HMI tags "ProNet Configuration"
   "PN_Mixinghead_Send" : Bool = PLC PN_Mixinghead.Send AT %DB1006.DBX4.0, 1 s
   "PN_Mixinghead_Mixinghead{0}_Digital_Address" : Int = PLC PN_Mixinghead.Mixinghead[0].Digital.Address AT %DB1006.DBW80, 1 s
      on ChangeValue: SetBit("PN_Mixinghead_Mixinghead{0}_Digital_Zeiten_Request"); SetBit("PN_Mixinghead_Mixinghead{0}_Digital_Zeiten_2_Request"); SetBit("PN_Mixinghead_Mixinghead{0}_Digital_GeneralParameters_Request")
   "PN_Mixinghead_Mixinghead{0}_Digital_Zeiten_Request" : Bool = PLC PN_Mixinghead.Mixinghead[0].Digital.Zeiten.Request AT %DB1006.DBX90.0, 1 s
   "PN_Mixinghead_Mixinghead{0}_Digital_Zeiten_Data_ÜberwachungszeitÖffnen" : Real = PLC PN_Mixinghead.Mixinghead[0].Digital.Zeiten.Data.ÜberwachungszeitÖffnen AT %DB1006.DBD92, 1 s
      on ChangeValue: SetBit("PN_Mixinghead_Mixinghead{0}_Digital_Zeiten_Request")
   "PN_Mixinghead_Mixinghead{0}_Digital_GeneralParameters_Data_MischkopfKanal" : Byte = PLC PN_Mixinghead.Mixinghead[0].Digital.GeneralParameters.Data.MischkopfKanal AT %DB1006.DBB89, 1 s
      on ChangeValue: SetBit("PN_Mixinghead_Mixinghead{0}_Digital_GeneralParameters_Request")
   "PN_Mixinghead_Mixinghead{0}_Digital_GeneralParameters_Request" : Bool = PLC PN_Mixinghead.Mixinghead[0].Digital.GeneralParameters.Request AT %DB1006.DBX84.0, 1 s
   "PN_Mixinghead_Mixinghead{0}_Digital_Active" : Bool = PLC PN_Mixinghead.Mixinghead[0].Digital.Active AT %DB1006.DBX82.0, 1 s
      on ChangeValue: SetBit("PN_Mixinghead_Mixinghead{0}_Digital_Zeiten_Request"); SetBit("PN_Mixinghead_Mixinghead{0}_Digital_Zeiten_2_Request"); SetBit("PN_Mixinghead_Mixinghead{0}_Digital_GeneralParameters_Request")
   "PN_Mixinghead_Mixinghead{0}_Digital_Zeiten_Data_ÜberwachungszeitSchließen" : Real = PLC PN_Mixinghead.Mixinghead[0].Digital.Zeiten.Data.ÜberwachungszeitSchließen AT %DB1006.DBD96, 1 s
      on ChangeValue: SetBit("PN_Mixinghead_Mixinghead{0}_Digital_Zeiten_Request")
   "PN_Mixinghead_Mixinghead{0}_Digital_Zeiten_Data_ErlaubtePrellzeit" : Real = PLC PN_Mixinghead.Mixinghead[0].Digital.Zeiten.Data.ErlaubtePrellzeit AT %DB1006.DBD100, 1 s
      on ChangeValue: SetBit("PN_Mixinghead_Mixinghead{0}_Digital_Zeiten_Request")
   "PN_Mixinghead_Mixinghead{0}_Digital_GeneralParameters_Data_Ventilausgang" : Byte = PLC PN_Mixinghead.Mixinghead[0].Digital.GeneralParameters.Data.Ventilausgang AT %DB1006.DBB88, 1 s
      on ChangeValue: SetBit("PN_Mixinghead_Mixinghead{0}_Digital_GeneralParameters_Request")
   "PN_Mixinghead_Mixinghead{0}_Digital_GeneralParameters_Data_EingangskanalMK_Ini" : Byte = PLC PN_Mixinghead.Mixinghead[0].Digital.GeneralParameters.Data.EingangskanalMK_Ini AT %DB1006.DBB86, 1 s
      on ChangeValue: SetBit("PN_Mixinghead_Mixinghead{0}_Digital_GeneralParameters_Request")
   "PN_Mixinghead_Mixinghead{0}_Digital_GeneralParameters_Data_EingangskanalFreigabe" : Byte = PLC PN_Mixinghead.Mixinghead[0].Digital.GeneralParameters.Data.EingangskanalFreigabe AT %DB1006.DBB87, 1 s
      on ChangeValue: SetBit("PN_Mixinghead_Mixinghead{0}_Digital_GeneralParameters_Request")
   "PN_Mixinghead_Mixinghead{0}_Digital_Zeiten_2_Request" : Bool = PLC PN_Mixinghead.Mixinghead[0].Digital.Zeiten_2.Request AT %DB1006.DBX104.0, 1 s
   "PN_Mixinghead_Mixinghead{0}_Digital_Zeiten_2_Data_Verzögerungszeit_HW_Freigabe" : Real = PLC PN_Mixinghead.Mixinghead[0].Digital.Zeiten_2.Data.Verzögerungszeit_HW_Freigabe AT %DB1006.DBD106, 1 s
      on ChangeValue: SetBit("PN_Mixinghead_Mixinghead{0}_Digital_Zeiten_2_Request")
   "PN_Mixinghead_SetIndex" : Int = PLC PN_Mixinghead.SetIndex AT %DB1006.DBW0, 1 s
   "PN_Mixinghead_Mixinghead{0}_ReinigungskolbenDigital_Active" : Bool = PLC PN_Mixinghead.Mixinghead[0].ReinigungskolbenDigital.Active AT %DB1006.DBX112.0, 1 s
      on ChangeValue: SetBit("PN_Mixinghead_Mixinghead{0}_ReinigungskolbenDigital_Zeiten_Request"); SetBit("PN_Mixinghead_Mixinghead{0}_ReinigungskolbenDigital_GeneralParameters_Request")
   "PN_Mixinghead_Mixinghead{0}_ReinigungskolbenDigital_GeneralParameters_Request" : Bool = PLC PN_Mixinghead.Mixinghead[0].ReinigungskolbenDigital.GeneralParameters.Request AT %DB1006.DBX114.0, 1 s
   "PN_Mixinghead_Mixinghead{0}_ReinigungskolbenDigital_GeneralParameters_Data_EingangskanalRK_Ini" : Byte = PLC PN_Mixinghead.Mixinghead[0].ReinigungskolbenDigital.GeneralParameters.Data.EingangskanalRK_Ini AT %DB1006.DBB116, 1 s
      on ChangeValue: SetBit("PN_Mixinghead_Mixinghead{0}_ReinigungskolbenDigital_GeneralParameters_Request")
   "PN_Mixinghead_Mixinghead{0}_ReinigungskolbenDigital_GeneralParameters_Data_AusgangRKVentil" : Byte = PLC PN_Mixinghead.Mixinghead[0].ReinigungskolbenDigital.GeneralParameters.Data.AusgangRKVentil AT %DB1006.DBB117, 1 s
      on ChangeValue: SetBit("PN_Mixinghead_Mixinghead{0}_ReinigungskolbenDigital_GeneralParameters_Request")
   "PN_Mixinghead_Mixinghead{0}_ReinigungskolbenDigital_GeneralParameters_Data_MischkopfKanal" : Byte = PLC PN_Mixinghead.Mixinghead[0].ReinigungskolbenDigital.GeneralParameters.Data.MischkopfKanal AT %DB1006.DBB118, 1 s
      on ChangeValue: SetBit("PN_Mixinghead_Mixinghead{0}_ReinigungskolbenDigital_GeneralParameters_Request")
   "PN_Mixinghead_Mixinghead{0}_ReinigungskolbenDigital_Address" : Int = PLC PN_Mixinghead.Mixinghead[0].ReinigungskolbenDigital.Address AT %DB1006.DBW110, 1 s
      on ChangeValue: SetBit("PN_Mixinghead_Mixinghead{0}_Digital_Zeiten_Request"); SetBit("PN_Mixinghead_Mixinghead{0}_Digital_Zeiten_2_Request"); SetBit("PN_Mixinghead_Mixinghead{0}_Digital_GeneralParameters_Request")
   "PN_Mixinghead_Mixinghead{0}_ReinigungskolbenDigital_Zeiten_Data_ÜberwachungszeitVorfahren" : Real = PLC PN_Mixinghead.Mixinghead[0].ReinigungskolbenDigital.Zeiten.Data.ÜberwachungszeitVorfahren AT %DB1006.DBD122, 1 s
      on ChangeValue: SetBit("PN_Mixinghead_Mixinghead{0}_ReinigungskolbenDigital_Zeiten_Request")
   "PN_Mixinghead_Mixinghead{0}_ReinigungskolbenDigital_Zeiten_Data_ÜberwachungszeitRückfahren" : Real = PLC PN_Mixinghead.Mixinghead[0].ReinigungskolbenDigital.Zeiten.Data.ÜberwachungszeitRückfahren AT %DB1006.DBD126, 1 s
      on ChangeValue: SetBit("PN_Mixinghead_Mixinghead{0}_ReinigungskolbenDigital_Zeiten_Request")
   "PN_Mixinghead_Mixinghead{0}_ReinigungskolbenDigital_Zeiten_Request" : Bool = PLC PN_Mixinghead.Mixinghead[0].ReinigungskolbenDigital.Zeiten.Request AT %DB1006.DBX120.0, 1 s
   "PN_Mixinghead_Mixinghead{0}_ReinigungskolbenDigital_Zeiten_Data_ErlaubtePrellzeit" : Real = PLC PN_Mixinghead.Mixinghead[0].ReinigungskolbenDigital.Zeiten.Data.ErlaubtePrellzeit AT %DB1006.DBD130, 1 s
      on ChangeValue: SetBit("PN_Mixinghead_Mixinghead{0}_ReinigungskolbenDigital_Zeiten_Request")
   "PN_Mixinghead_Mixinghead{0}_ReinigungskolbenDigital_Zeiten_Data_WartezeitVorne" : Real = PLC PN_Mixinghead.Mixinghead[0].ReinigungskolbenDigital.Zeiten.Data.WartezeitVorne AT %DB1006.DBD134, 1 s
      on ChangeValue: SetBit("PN_Mixinghead_Mixinghead{0}_ReinigungskolbenDigital_Zeiten_Request")
   "PN_Mixinghead_Mixinghead{0}_ReinigungskolbenDigital_Zeiten_Data_VerzögerungNachSchuss" : Real = PLC PN_Mixinghead.Mixinghead[0].ReinigungskolbenDigital.Zeiten.Data.VerzögerungNachSchuss AT %DB1006.DBD138, 1 s
      on ChangeValue: SetBit("PN_Mixinghead_Mixinghead{0}_ReinigungskolbenDigital_Zeiten_Request")
   "PN_AI_Send" : Bool = PLC PN_AI.Send AT %DB1002.DBX4.0, 1 s
   "PN_AI_Module{0}_AI8_Address" : Int = PLC PN_AI.Module[0].AI8.Address AT %DB1002.DBW6, 1 s
      on ChangeValue: SetBit("PN_AI_Send"); SetBit("PN_AI_Module{0}_AI8_X14_0_Request")
   "PN_AI_Module{0}_AI8_Active" : Bool = PLC PN_AI.Module[0].AI8.Active AT %DB1002.DBX8.0, 1 s
      on ChangeValue: SetBit("PN_AI_Send"); SetBit("PN_AI_Module{0}_AI8_X14_0_Request")
   "PN_AI_Module{0}_AI8_X14_0_Data_Data[1]_Betriebsart" : Byte = PLC PN_AI.Module[0].AI8.X14_0.Data."Data[1]".Betriebsart AT %DB1002.DBB12, 1 s
      on ChangeValue: SetBit("PN_AI_Send"); SetBit("PN_AI_Module{0}_AI8_X14_0_Request")
   "PN_AI_Module{0}_AI8_X14_0_Data_Data[2]_Betriebsart" : Byte = PLC PN_AI.Module[0].AI8.X14_0.Data."Data[2]".Betriebsart AT %DB1002.DBB20, 1 s
      on ChangeValue: SetBit("PN_AI_Send"); SetBit("PN_AI_Module{0}_AI8_X14_0_Request")
   "PN_AI_Module{0}_AI8_X14_0_Data_Data[1]_Bereichsuntergrenze" : Int = PLC PN_AI.Module[0].AI8.X14_0.Data."Data[1]".Bereichsuntergrenze AT %DB1002.DBW16, 1 s
      on ChangeValue: SetBit("PN_AI_Send"); SetBit("PN_AI_Module{0}_AI8_X14_0_Request")
   "PN_AI_Module{0}_AI8_X14_0_Data_Data[1]_Bereichsobergrenze" : Int = PLC PN_AI.Module[0].AI8.X14_0.Data."Data[1]".Bereichsobergrenze AT %DB1002.DBW14, 1 s
      on ChangeValue: SetBit("PN_AI_Send"); SetBit("PN_AI_Module{0}_AI8_X14_0_Request")
   "PN_AI_Module{0}_AI8_X14_0_Data_Data[1]_Mittelwertzeit" : Int = PLC PN_AI.Module[0].AI8.X14_0.Data."Data[1]".Mittelwertzeit AT %DB1002.DBW18, 1 s
      on ChangeValue: SetBit("PN_AI_Send"); SetBit("PN_AI_Module{0}_AI8_X14_0_Request")
   "PN_AI_Module{0}_AI8_X14_0_Data_Data[2]_Bereichsobergrenze" : Int = PLC PN_AI.Module[0].AI8.X14_0.Data."Data[2]".Bereichsobergrenze AT %DB1002.DBW22, 1 s
      on ChangeValue: SetBit("PN_AI_Send"); SetBit("PN_AI_Module{0}_AI8_X14_0_Request")
   "PN_AI_Module{0}_AI8_X14_0_Data_Data[2]_Bereichsuntergrenze" : Int = PLC PN_AI.Module[0].AI8.X14_0.Data."Data[2]".Bereichsuntergrenze AT %DB1002.DBW24, 1 s
      on ChangeValue: SetBit("PN_AI_Send"); SetBit("PN_AI_Module{0}_AI8_X14_0_Request")
   "PN_AI_Module{0}_AI8_X14_0_Data_Data[2]_Mittelwertzeit" : Int = PLC PN_AI.Module[0].AI8.X14_0.Data."Data[2]".Mittelwertzeit AT %DB1002.DBW26, 1 s
      on ChangeValue: SetBit("PN_AI_Send"); SetBit("PN_AI_Module{0}_AI8_X14_0_Request")
   "PN_AI_Module{0}_AI8_X14_0_Data_Data[3]_Betriebsart" : Byte = PLC PN_AI.Module[0].AI8.X14_0.Data."Data[3]".Betriebsart AT %DB1002.DBB28, 1 s
      on ChangeValue: SetBit("PN_AI_Send"); SetBit("PN_AI_Module{0}_AI8_X14_0_Request")
   "PN_Mixinghead_Mixinghead{0}_DüseBypass{6}_Zeiten_Request" : Bool = PLC PN_Mixinghead.Mixinghead[0].DüseBypass[6].Zeiten.Request AT %DB1006.DBX458.0, 1 s
      on ChangeValue: SetBit("PN_AI_Send"); SetBit("PN_AI_Module{0}_AI8_X14_0_Request")
   "PN_AI_Module{0}_AI8_X14_0_Data_Data[3]_Bereichsuntergrenze" : Int = PLC PN_AI.Module[0].AI8.X14_0.Data."Data[3]".Bereichsuntergrenze AT %DB1002.DBW32, 1 s
      on ChangeValue: SetBit("PN_AI_Send"); SetBit("PN_AI_Module{0}_AI8_X14_0_Request")
   "PN_AI_Module{0}_AI8_X14_0_Data_Data[3]_Mittelwertzeit" : Int = PLC PN_AI.Module[0].AI8.X14_0.Data."Data[3]".Mittelwertzeit AT %DB1002.DBW34, 1 s
      on ChangeValue: SetBit("PN_AI_Send"); SetBit("PN_AI_Module{0}_AI8_X14_0_Request")
   "PN_AI_Module{0}_AI8_X14_0_Data_Data[4]_Betriebsart" : Byte = PLC PN_AI.Module[0].AI8.X14_0.Data."Data[4]".Betriebsart AT %DB1002.DBB36, 1 s
      on ChangeValue: SetBit("PN_AI_Send"); SetBit("PN_AI_Module{0}_AI8_X14_0_Request")
   "PN_AI_Module{0}_AI8_X14_0_Data_Data[4]_Bereichsobergrenze" : Int = PLC PN_AI.Module[0].AI8.X14_0.Data."Data[4]".Bereichsobergrenze AT %DB1002.DBW38, 1 s
      on ChangeValue: SetBit("PN_AI_Send"); SetBit("PN_AI_Module{0}_AI8_X14_0_Request")
   "PN_AI_Module{0}_AI8_X14_0_Data_Data[4]_Bereichsuntergrenze" : Int = PLC PN_AI.Module[0].AI8.X14_0.Data."Data[4]".Bereichsuntergrenze AT %DB1002.DBW40, 1 s
      on ChangeValue: SetBit("PN_AI_Send"); SetBit("PN_AI_Module{0}_AI8_X14_0_Request")
   "PN_AI_Module{0}_AI8_X14_0_Data_Data[4]_Mittelwertzeit" : Int = PLC PN_AI.Module[0].AI8.X14_0.Data."Data[4]".Mittelwertzeit AT %DB1002.DBW42, 1 s
      on ChangeValue: SetBit("PN_AI_Send"); SetBit("PN_AI_Module{0}_AI8_X14_0_Request")
   "PN_AI_Module{0}_AI8_X14_0_Data_Data[5]_Betriebsart" : Byte = PLC PN_AI.Module[0].AI8.X14_0.Data."Data[5]".Betriebsart AT %DB1002.DBB44, 1 s
      on ChangeValue: SetBit("PN_AI_Send"); SetBit("PN_AI_Module{0}_AI8_X14_0_Request")
   "PN_AI_Module{0}_AI8_X14_0_Data_Data[5]_Bereichsobergrenze" : Int = PLC PN_AI.Module[0].AI8.X14_0.Data."Data[5]".Bereichsobergrenze AT %DB1002.DBW46, 1 s
      on ChangeValue: SetBit("PN_AI_Send"); SetBit("PN_AI_Module{0}_AI8_X14_0_Request")
   "PN_AI_Module{0}_AI8_X14_0_Data_Data[5]_Bereichsuntergrenze" : Int = PLC PN_AI.Module[0].AI8.X14_0.Data."Data[5]".Bereichsuntergrenze AT %DB1002.DBW48, 1 s
      on ChangeValue: SetBit("PN_AI_Send"); SetBit("PN_AI_Module{0}_AI8_X14_0_Request")
   "PN_AI_Module{0}_AI8_X14_0_Data_Data[5]_Mittelwertzeit" : Int = PLC PN_AI.Module[0].AI8.X14_0.Data."Data[5]".Mittelwertzeit AT %DB1002.DBW50, 1 s
      on ChangeValue: SetBit("PN_AI_Send"); SetBit("PN_AI_Module{0}_AI8_X14_0_Request")
   "PN_AI_Module{0}_AI8_X14_0_Data_Data[6]_Betriebsart" : Byte = PLC PN_AI.Module[0].AI8.X14_0.Data."Data[6]".Betriebsart AT %DB1002.DBB52, 1 s
      on ChangeValue: SetBit("PN_AI_Send"); SetBit("PN_AI_Module{0}_AI8_X14_0_Request")
   "PN_AI_Module{0}_AI8_X14_0_Data_Data[6]_Bereichsobergrenze" : Int = PLC PN_AI.Module[0].AI8.X14_0.Data."Data[6]".Bereichsobergrenze AT %DB1002.DBW54, 1 s
      on ChangeValue: SetBit("PN_AI_Send"); SetBit("PN_AI_Module{0}_AI8_X14_0_Request")
   "PN_AI_Module{0}_AI8_X14_0_Data_Data[6]_Bereichsuntergrenze" : Int = PLC PN_AI.Module[0].AI8.X14_0.Data."Data[6]".Bereichsuntergrenze AT %DB1002.DBW56, 1 s
      on ChangeValue: SetBit("PN_AI_Send"); SetBit("PN_AI_Module{0}_AI8_X14_0_Request")
   "PN_AI_Module{0}_AI8_X14_0_Data_Data[6]_Mittelwertzeit" : Int = PLC PN_AI.Module[0].AI8.X14_0.Data."Data[6]".Mittelwertzeit AT %DB1002.DBW58, 1 s
      on ChangeValue: SetBit("PN_AI_Send"); SetBit("PN_AI_Module{0}_AI8_X14_0_Request")
   "PN_AI_Module{0}_AI8_X14_0_Data_Data[7]_Betriebsart" : Byte = PLC PN_AI.Module[0].AI8.X14_0.Data."Data[7]".Betriebsart AT %DB1002.DBB60, 1 s
      on ChangeValue: SetBit("PN_AI_Send"); SetBit("PN_AI_Module{0}_AI8_X14_0_Request")
   "PN_AI_Module{0}_AI8_X14_0_Data_Data[7]_Bereichsobergrenze" : Int = PLC PN_AI.Module[0].AI8.X14_0.Data."Data[7]".Bereichsobergrenze AT %DB1002.DBW62, 1 s
      on ChangeValue: SetBit("PN_AI_Send"); SetBit("PN_AI_Module{0}_AI8_X14_0_Request")
   "PN_AI_Module{0}_AI8_X14_0_Data_Data[7]_Bereichsuntergrenze" : Int = PLC PN_AI.Module[0].AI8.X14_0.Data."Data[7]".Bereichsuntergrenze AT %DB1002.DBW64, 1 s
      on ChangeValue: SetBit("PN_AI_Send"); SetBit("PN_AI_Module{0}_AI8_X14_0_Request")
   "PN_AI_Module{0}_AI8_X14_0_Data_Data[7]_Mittelwertzeit" : Int = PLC PN_AI.Module[0].AI8.X14_0.Data."Data[7]".Mittelwertzeit AT %DB1002.DBW66, 1 s
      on ChangeValue: SetBit("PN_AI_Send"); SetBit("PN_AI_Module{0}_AI8_X14_0_Request")
   "PN_AI_Module{0}_AI8_X14_0_Data_Data[8]_Betriebsart" : Byte = PLC PN_AI.Module[0].AI8.X14_0.Data."Data[8]".Betriebsart AT %DB1002.DBB68, 1 s
      on ChangeValue: SetBit("PN_AI_Send"); SetBit("PN_AI_Module{0}_AI8_X14_0_Request")
   "PN_AI_Module{0}_AI8_X14_0_Data_Data[8]_Bereichsobergrenze" : Int = PLC PN_AI.Module[0].AI8.X14_0.Data."Data[8]".Bereichsobergrenze AT %DB1002.DBW70, 1 s
      on ChangeValue: SetBit("PN_AI_Send"); SetBit("PN_AI_Module{0}_AI8_X14_0_Request")
   "PN_AI_Module{0}_AI8_X14_0_Data_Data[8]_Bereichsuntergrenze" : Int = PLC PN_AI.Module[0].AI8.X14_0.Data."Data[8]".Bereichsuntergrenze AT %DB1002.DBW72, 1 s
      on ChangeValue: SetBit("PN_AI_Send"); SetBit("PN_AI_Module{0}_AI8_X14_0_Request")
   "PN_AI_Module{0}_AI8_X14_0_Data_Data[8]_Mittelwertzeit" : Int = PLC PN_AI.Module[0].AI8.X14_0.Data."Data[8]".Mittelwertzeit AT %DB1002.DBW74, 1 s
      on ChangeValue: SetBit("PN_AI_Send"); SetBit("PN_AI_Module{0}_AI8_X14_0_Request")
   "PN_AI_Module{0}_AI8_X14_0_Request" : Bool = PLC PN_AI.Module[0].AI8.X14_0.Request AT %DB1002.DBX10.0, 1 s
   "PN_AI_SetIndex" : Int = PLC PN_AI.SetIndex AT %DB1002.DBW0, 1 s
      on ChangeValue: SetBit("PN_AI_Send")
   "PN_AI_Module{0}_AIResistive_8_Address" : Int = PLC PN_AI.Module[0].AIResistive_8.Address AT %DB1002.DBW76, 1 s
      on ChangeValue: SetBit("PN_AI_Send"); SetBit("PN_AI_Module{0}_AIResistive_8_TemperatureInput_Request")
   "PN_AI_Module{0}_AIResistive_8_TemperatureInput_Request" : Bool = PLC PN_AI.Module[0].AIResistive_8.TemperatureInput.Request AT %DB1002.DBX80.0, 1 s
      on ChangeValue: SetBit("PN_AI_Send")
   "PN_AI_Module{0}_AIResistive_8_Active" : Bool = PLC PN_AI.Module[0].AIResistive_8.Active AT %DB1002.DBX78.0, 1 s
      on ChangeValue: SetBit("PN_AI_Send")
   "PN_AI_Module{0}_AIResistive_8_TemperatureInput_Data{1}_Mittelwertzeit" : Int = PLC PN_AI.Module[0].AIResistive_8.TemperatureInput.Data[1].Mittelwertzeit AT %DB1002.DBW82, 1 s
      on ChangeValue: SetBit("PN_AI_Send"); SetBit("PN_AI_Module{0}_AIResistive_8_TemperatureInput_Request")
   "PN_AI_Module{0}_AIResistive_8_TemperatureInput_Data{1}_ErsatzwertDrahtbruch" : Int = PLC PN_AI.Module[0].AIResistive_8.TemperatureInput.Data[1].ErsatzwertDrahtbruch AT %DB1002.DBW84, 1 s
      on ChangeValue: SetBit("PN_AI_Send"); SetBit("PN_AI_Module{0}_AIResistive_8_TemperatureInput_Request")
   "PN_AI_Module{0}_AIResistive_8_TemperatureInput_Data{1}_Einheit" : Byte = PLC PN_AI.Module[0].AIResistive_8.TemperatureInput.Data[1].Einheit AT %DB1002.DBB86, 1 s
      on ChangeValue: SetBit("PN_AI_Send"); SetBit("PN_AI_Module{0}_AIResistive_8_TemperatureInput_Request")
   "PN_AI_Module{0}_AIResistive_8_TemperatureInput_Data{2}_Mittelwertzeit" : Int = PLC PN_AI.Module[0].AIResistive_8.TemperatureInput.Data[2].Mittelwertzeit AT %DB1002.DBW88, 1 s
      on ChangeValue: SetBit("PN_AI_Send"); SetBit("PN_AI_Module{0}_AIResistive_8_TemperatureInput_Request")
   "PN_AI_Module{0}_AIResistive_8_TemperatureInput_Data{2}_ErsatzwertDrahtbruch" : Int = PLC PN_AI.Module[0].AIResistive_8.TemperatureInput.Data[2].ErsatzwertDrahtbruch AT %DB1002.DBW90, 1 s
      on ChangeValue: SetBit("PN_AI_Send"); SetBit("PN_AI_Module{0}_AIResistive_8_TemperatureInput_Request")
   "PN_AI_Module{0}_AIResistive_8_TemperatureInput_Data{2}_Einheit" : Byte = PLC PN_AI.Module[0].AIResistive_8.TemperatureInput.Data[2].Einheit AT %DB1002.DBB92, 1 s
      on ChangeValue: SetBit("PN_AI_Send"); SetBit("PN_AI_Module{0}_AIResistive_8_TemperatureInput_Request")
   "PN_AI_Module{0}_AIResistive_8_TemperatureInput_Data{3}_Mittelwertzeit" : Int = PLC PN_AI.Module[0].AIResistive_8.TemperatureInput.Data[3].Mittelwertzeit AT %DB1002.DBW94, 1 s
      on ChangeValue: SetBit("PN_AI_Send"); SetBit("PN_AI_Module{0}_AIResistive_8_TemperatureInput_Request")
   "PN_AI_Module{0}_AIResistive_8_TemperatureInput_Data{3}_ErsatzwertDrahtbruch" : Int = PLC PN_AI.Module[0].AIResistive_8.TemperatureInput.Data[3].ErsatzwertDrahtbruch AT %DB1002.DBW96, 1 s
      on ChangeValue: SetBit("PN_AI_Send"); SetBit("PN_AI_Module{0}_AIResistive_8_TemperatureInput_Request")
   "PN_AI_Module{0}_AIResistive_8_TemperatureInput_Data{3}_Einheit" : Byte = PLC PN_AI.Module[0].AIResistive_8.TemperatureInput.Data[3].Einheit AT %DB1002.DBB98, 1 s
      on ChangeValue: SetBit("PN_AI_Send"); SetBit("PN_AI_Module{0}_AIResistive_8_TemperatureInput_Request")
   "PN_AI_Module{0}_AIResistive_8_TemperatureInput_Data{4}_Mittelwertzeit" : Int = PLC PN_AI.Module[0].AIResistive_8.TemperatureInput.Data[4].Mittelwertzeit AT %DB1002.DBW100, 1 s
      on ChangeValue: SetBit("PN_AI_Send"); SetBit("PN_AI_Module{0}_AIResistive_8_TemperatureInput_Request")
   "PN_AI_Module{0}_AIResistive_8_TemperatureInput_Data{4}_ErsatzwertDrahtbruch" : Int = PLC PN_AI.Module[0].AIResistive_8.TemperatureInput.Data[4].ErsatzwertDrahtbruch AT %DB1002.DBW102, 1 s
      on ChangeValue: SetBit("PN_AI_Send"); SetBit("PN_AI_Module{0}_AIResistive_8_TemperatureInput_Request")
   "PN_AI_Module{0}_AIResistive_8_TemperatureInput_Data{4}_Einheit" : Byte = PLC PN_AI.Module[0].AIResistive_8.TemperatureInput.Data[4].Einheit AT %DB1002.DBB104, 1 s
      on ChangeValue: SetBit("PN_AI_Send"); SetBit("PN_AI_Module{0}_AIResistive_8_TemperatureInput_Request")
   "PN_AI_Module{0}_AIResistive_8_TemperatureInput_Data{5}_Mittelwertzeit" : Int = PLC PN_AI.Module[0].AIResistive_8.TemperatureInput.Data[5].Mittelwertzeit AT %DB1002.DBW106, 1 s
      on ChangeValue: SetBit("PN_AI_Send"); SetBit("PN_AI_Module{0}_AIResistive_8_TemperatureInput_Request")
   "PN_AI_Module{0}_AIResistive_8_TemperatureInput_Data{5}_ErsatzwertDrahtbruch" : Int = PLC PN_AI.Module[0].AIResistive_8.TemperatureInput.Data[5].ErsatzwertDrahtbruch AT %DB1002.DBW108, 1 s
      on ChangeValue: SetBit("PN_AI_Send"); SetBit("PN_AI_Module{0}_AIResistive_8_TemperatureInput_Request")
   "PN_AI_Module{0}_AIResistive_8_TemperatureInput_Data{5}_Einheit" : Byte = PLC PN_AI.Module[0].AIResistive_8.TemperatureInput.Data[5].Einheit AT %DB1002.DBB110, 1 s
      on ChangeValue: SetBit("PN_AI_Send"); SetBit("PN_AI_Module{0}_AIResistive_8_TemperatureInput_Request")
   "PN_AI_Module{0}_AIResistive_8_TemperatureInput_Data{6}_Mittelwertzeit" : Int = PLC PN_AI.Module[0].AIResistive_8.TemperatureInput.Data[6].Mittelwertzeit AT %DB1002.DBW112, 1 s
      on ChangeValue: SetBit("PN_AI_Send"); SetBit("PN_AI_Module{0}_AIResistive_8_TemperatureInput_Request")
   "PN_AI_Module{0}_AIResistive_8_TemperatureInput_Data{6}_ErsatzwertDrahtbruch" : Int = PLC PN_AI.Module[0].AIResistive_8.TemperatureInput.Data[6].ErsatzwertDrahtbruch AT %DB1002.DBW114, 1 s
      on ChangeValue: SetBit("PN_AI_Send"); SetBit("PN_AI_Module{0}_AIResistive_8_TemperatureInput_Request")
   "PN_AI_Module{0}_AIResistive_8_TemperatureInput_Data{6}_Einheit" : Byte = PLC PN_AI.Module[0].AIResistive_8.TemperatureInput.Data[6].Einheit AT %DB1002.DBB116, 1 s
      on ChangeValue: SetBit("PN_AI_Send"); SetBit("PN_AI_Module{0}_AIResistive_8_TemperatureInput_Request")
   "PN_AI_Module{0}_AIResistive_8_TemperatureInput_Data{7}_Mittelwertzeit" : Int = PLC PN_AI.Module[0].AIResistive_8.TemperatureInput.Data[7].Mittelwertzeit AT %DB1002.DBW118, 1 s
      on ChangeValue: SetBit("PN_AI_Send"); SetBit("PN_AI_Module{0}_AIResistive_8_TemperatureInput_Request")
   "PN_AI_Module{0}_AIResistive_8_TemperatureInput_Data{7}_ErsatzwertDrahtbruch" : Int = PLC PN_AI.Module[0].AIResistive_8.TemperatureInput.Data[7].ErsatzwertDrahtbruch AT %DB1002.DBW120, 1 s
      on ChangeValue: SetBit("PN_AI_Send"); SetBit("PN_AI_Module{0}_AIResistive_8_TemperatureInput_Request")
   "PN_AI_Module{0}_AIResistive_8_TemperatureInput_Data{7}_Einheit" : Byte = PLC PN_AI.Module[0].AIResistive_8.TemperatureInput.Data[7].Einheit AT %DB1002.DBB122, 1 s
      on ChangeValue: SetBit("PN_AI_Send"); SetBit("PN_AI_Module{0}_AIResistive_8_TemperatureInput_Request")
   "PN_AI_Module{0}_AIResistive_8_TemperatureInput_Data{8}_Mittelwertzeit" : Int = PLC PN_AI.Module[0].AIResistive_8.TemperatureInput.Data[8].Mittelwertzeit AT %DB1002.DBW124, 1 s
      on ChangeValue: SetBit("PN_AI_Send"); SetBit("PN_AI_Module{0}_AIResistive_8_TemperatureInput_Request")
   "PN_AI_Module{0}_AIResistive_8_TemperatureInput_Data{8}_ErsatzwertDrahtbruch" : Int = PLC PN_AI.Module[0].AIResistive_8.TemperatureInput.Data[8].ErsatzwertDrahtbruch AT %DB1002.DBW126, 1 s
      on ChangeValue: SetBit("PN_AI_Send"); SetBit("PN_AI_Module{0}_AIResistive_8_TemperatureInput_Request")
   "PN_AI_Module{0}_AIResistive_8_TemperatureInput_Data{8}_Einheit" : Byte = PLC PN_AI.Module[0].AIResistive_8.TemperatureInput.Data[8].Einheit AT %DB1002.DBB128, 1 s
      on ChangeValue: SetBit("PN_AI_Send"); SetBit("PN_AI_Module{0}_AIResistive_8_TemperatureInput_Request")
   "PN_FlowRate_Component{0}_FlowC_F_Address" : Int = PLC PN_FlowRate.Component[0].FlowC_F.Address AT %DB1003.DBW54, 1 s
      on ChangeValue: SetBit("PN_FlowRate_Send")
   "PN_FlowRate_Component{0}_FlowC_F_Active" : Bool = PLC PN_FlowRate.Component[0].FlowC_F.Active AT %DB1003.DBX56.0, 1 s
      on ChangeValue: SetBit("PN_FlowRate_Component{0}_FlowC_F_Hardware_Request"); SetBit("PN_FlowRate_Component{0}_FlowC_F_GeneralParameters_Request"); SetBit("PN_FlowRate_Component{0}_FlowC_F_Grenzen_Request"); SetBit("PN_FlowRate_Component{0}_FlowC_F_SkalierungAI_Request")
   "PN_FlowRate_Component{0}_FlowC_F_Hardware_Request" : Bool = PLC PN_FlowRate.Component[0].FlowC_F.Hardware.Request AT %DB1003.DBX88.0, 1 s
   "PN_FlowRate_Component{0}_FlowC_F_GeneralParameters_Request" : Bool = PLC PN_FlowRate.Component[0].FlowC_F.GeneralParameters.Request AT %DB1003.DBX100.0, 1 s
   "PN_FlowRate_Component{0}_FlowC_F_Grenzen_Request" : Bool = PLC PN_FlowRate.Component[0].FlowC_F.Grenzen.Request AT %DB1003.DBX118.0, 1 s
   "PN_FlowRate_Component{0}_FlowC_F_SkalierungAI_Request" : Bool = PLC PN_FlowRate.Component[0].FlowC_F.SkalierungAI.Request AT %DB1003.DBX136.0, 1 s
   "PN_FlowRate_Send" : Bool = PLC PN_FlowRate.Send AT %DB1003.DBX4.0, 1 s
   "PN_FlowRate_Component{0}_FlowC_F_SkalierungAI_Data_Bereichsobergrenze" : Real = PLC PN_FlowRate.Component[0].FlowC_F.SkalierungAI.Data.Bereichsobergrenze AT %DB1003.DBD138, 1 s
      on ChangeValue: SetBit("PN_FlowRate_Send"); SetBit("PN_FlowRate_Component{0}_FlowC_F_SkalierungAI_Request")
   "PN_FlowRate_Component{0}_FlowC_F_SkalierungAI_Data_Bereichsuntergrenze" : Real = PLC PN_FlowRate.Component[0].FlowC_F.SkalierungAI.Data.Bereichsuntergrenze AT %DB1003.DBD142, 1 s
      on ChangeValue: SetBit("PN_FlowRate_Send"); SetBit("PN_FlowRate_Component{0}_FlowC_F_SkalierungAI_Request")
   "PN_FlowRate_Component{0}_FlowC_F_SkalierungAI_Data_Mittelwertzeit" : Real = PLC PN_FlowRate.Component[0].FlowC_F.SkalierungAI.Data.Mittelwertzeit AT %DB1003.DBD146, 1 s
      on ChangeValue: SetBit("PN_FlowRate_Send"); SetBit("PN_FlowRate_Component{0}_FlowC_F_SkalierungAI_Request")
   "PN_FlowRate_SetIndex" : Int = PLC PN_FlowRate.SetIndex AT %DB1003.DBW0, 1 s
      on ChangeValue: SetBit("PN_FlowRate_Send")
   "PN_FlowRate_Component{0}_FlowC_F_GeneralParameters_Data_Filterzeit" : Real = PLC PN_FlowRate.Component[0].FlowC_F.GeneralParameters.Data.Filterzeit AT %DB1003.DBD114, 1 s
      on ChangeValue: SetBit("PN_FlowRate_Send"); SetBit("PN_FlowRate_Component{0}_FlowC_F_GeneralParameters_Request")
   "PN_FlowRate_Component{0}_FlowC_F_GeneralParameters_Data_Kalibrierfaktor" : Real = PLC PN_FlowRate.Component[0].FlowC_F.GeneralParameters.Data.Kalibrierfaktor AT %DB1003.DBD102, 1 s
      on ChangeValue: SetBit("PN_FlowRate_Send"); SetBit("PN_FlowRate_Component{0}_FlowC_F_GeneralParameters_Request")
   "PN_FlowRate_Component{0}_FlowC_F_GeneralParameters_Data_MaxDurchfluss" : Real = PLC PN_FlowRate.Component[0].FlowC_F.GeneralParameters.Data.MaxDurchfluss AT %DB1003.DBD106, 1 s
      on ChangeValue: SetBit("PN_FlowRate_Send"); SetBit("PN_FlowRate_Component{0}_FlowC_F_GeneralParameters_Request")
   "PN_FlowRate_Component{0}_FlowC_F_GeneralParameters_Data_Nachstellzeit" : Real = PLC PN_FlowRate.Component[0].FlowC_F.GeneralParameters.Data.Nachstellzeit AT %DB1003.DBD110, 1 s
      on ChangeValue: SetBit("PN_FlowRate_Send"); SetBit("PN_FlowRate_Component{0}_FlowC_F_GeneralParameters_Request")
   "PN_FlowRate_Component{0}_FlowC_F_Grenzen_Data_ObergrenzeStellgröße" : Real = PLC PN_FlowRate.Component[0].FlowC_F.Grenzen.Data.ObergrenzeStellgröße AT %DB1003.DBD120, 1 s
      on ChangeValue: SetBit("PN_FlowRate_Send"); SetBit("PN_FlowRate_Component{0}_FlowC_F_Grenzen_Request")
   "PN_FlowRate_Component{0}_FlowC_F_Grenzen_Data_UntergrenzeStellgröße" : Real = PLC PN_FlowRate.Component[0].FlowC_F.Grenzen.Data.UntergrenzeStellgröße AT %DB1003.DBD124, 1 s
      on ChangeValue: SetBit("PN_FlowRate_Send"); SetBit("PN_FlowRate_Component{0}_FlowC_F_Grenzen_Request")
   "PN_FlowRate_Component{0}_FlowC_F_Grenzen_Data_VerzögerungAlarmObergrenze" : Real = PLC PN_FlowRate.Component[0].FlowC_F.Grenzen.Data.VerzögerungAlarmObergrenze AT %DB1003.DBD128, 1 s
      on ChangeValue: SetBit("PN_FlowRate_Send"); SetBit("PN_FlowRate_Component{0}_FlowC_F_Grenzen_Request")
   "PN_FlowRate_Component{0}_FlowC_F_Grenzen_Data_VerzögerungAlarmUntergrenze" : Real = PLC PN_FlowRate.Component[0].FlowC_F.Grenzen.Data.VerzögerungAlarmUntergrenze AT %DB1003.DBD132, 1 s
      on ChangeValue: SetBit("PN_FlowRate_Send"); SetBit("PN_FlowRate_Component{0}_FlowC_F_Grenzen_Request")
   "PN_Mixinghead_Mixinghead{0}_DüseBypass{1}_Address" : Int = PLC PN_Mixinghead.Mixinghead[0].DüseBypass[1].Address AT %DB1006.DBW278, 1 s
      on ChangeValue: SetBit("PN_Mixinghead_Send"); SetBit("PN_Mixinghead_Mixinghead{0}_DüseBypass{1}_Channel_Request"); SetBit("PN_Mixinghead_Mixinghead{0}_DüseBypass{1}_Zeiten_Request")
   "PN_Mixinghead_Mixinghead{0}_DüseBypass{1}_Active" : Bool = PLC PN_Mixinghead.Mixinghead[0].DüseBypass[1].Active AT %DB1006.DBX280.0, 1 s
      on ChangeValue: SetBit("PN_Mixinghead_Send"); SetBit("PN_Mixinghead_Mixinghead{0}_DüseBypass{1}_Channel_Request"); SetBit("PN_Mixinghead_Mixinghead{0}_DüseBypass{1}_Zeiten_Request")
   "PN_Mixinghead_Mixinghead{0}_DüseBypass{2}_Address" : Int = PLC PN_Mixinghead.Mixinghead[0].DüseBypass[2].Address AT %DB1006.DBW312, 1 s
      on ChangeValue: SetBit("PN_Mixinghead_Send"); SetBit("PN_Mixinghead_Mixinghead{0}_DüseBypass{2}_Channel_Request"); SetBit("PN_Mixinghead_Mixinghead{0}_DüseBypass{2}_Zeiten_Request")
   "PN_Mixinghead_Mixinghead{0}_DüseBypass{2}_Active" : Bool = PLC PN_Mixinghead.Mixinghead[0].DüseBypass[2].Active AT %DB1006.DBX314.0, 1 s
      on ChangeValue: SetBit("PN_Mixinghead_Send"); SetBit("PN_Mixinghead_Mixinghead{0}_DüseBypass{2}_Channel_Request"); SetBit("PN_Mixinghead_Mixinghead{0}_DüseBypass{2}_Zeiten_Request")
   "PN_Mixinghead_Mixinghead{0}_DüseBypass{3}_Address" : Int = PLC PN_Mixinghead.Mixinghead[0].DüseBypass[3].Address AT %DB1006.DBW346, 1 s
      on ChangeValue: SetBit("PN_Mixinghead_Send"); SetBit("PN_Mixinghead_Mixinghead{0}_DüseBypass{3}_Channel_Request"); SetBit("PN_Mixinghead_Mixinghead{0}_DüseBypass{3}_Zeiten_Request")
   "PN_Mixinghead_Mixinghead{0}_DüseBypass{3}_Active" : Bool = PLC PN_Mixinghead.Mixinghead[0].DüseBypass[3].Active AT %DB1006.DBX348.0, 1 s
      on ChangeValue: SetBit("PN_Mixinghead_Send"); SetBit("PN_Mixinghead_Mixinghead{0}_DüseBypass{3}_Channel_Request"); SetBit("PN_Mixinghead_Mixinghead{0}_DüseBypass{3}_Zeiten_Request")
   "PN_Mixinghead_Mixinghead{0}_DüseBypass{4}_Address" : Int = PLC PN_Mixinghead.Mixinghead[0].DüseBypass[4].Address AT %DB1006.DBW380, 1 s
      on ChangeValue: SetBit("PN_Mixinghead_Send"); SetBit("PN_Mixinghead_Mixinghead{0}_DüseBypass{4}_Channel_Request"); SetBit("PN_Mixinghead_Mixinghead{0}_DüseBypass{4}_Zeiten_Request")
   "PN_Mixinghead_Mixinghead{0}_DüseBypass{4}_Active" : Bool = PLC PN_Mixinghead.Mixinghead[0].DüseBypass[4].Active AT %DB1006.DBX382.0, 1 s
      on ChangeValue: SetBit("PN_Mixinghead_Send"); SetBit("PN_Mixinghead_Mixinghead{0}_DüseBypass{4}_Channel_Request"); SetBit("PN_Mixinghead_Mixinghead{0}_DüseBypass{4}_Zeiten_Request")
   "PN_Mixinghead_Mixinghead{0}_DüseBypass{5}_Address" : Int = PLC PN_Mixinghead.Mixinghead[0].DüseBypass[5].Address AT %DB1006.DBW414, 1 s
      on ChangeValue: SetBit("PN_Mixinghead_Send"); SetBit("PN_Mixinghead_Mixinghead{0}_DüseBypass{5}_Channel_Request"); SetBit("PN_Mixinghead_Mixinghead{0}_DüseBypass{5}_Zeiten_Request")
   "PN_Mixinghead_Mixinghead{0}_DüseBypass{5}_Active" : Bool = PLC PN_Mixinghead.Mixinghead[0].DüseBypass[5].Active AT %DB1006.DBX416.0, 1 s
      on ChangeValue: SetBit("PN_Mixinghead_Send"); SetBit("PN_Mixinghead_Mixinghead{0}_DüseBypass{5}_Channel_Request"); SetBit("PN_Mixinghead_Mixinghead{0}_DüseBypass{5}_Zeiten_Request")
   "PN_Mixinghead_Mixinghead{0}_DüseBypass{6}_Address" : Int = PLC PN_Mixinghead.Mixinghead[0].DüseBypass[6].Address AT %DB1006.DBW448, 1 s
      on ChangeValue: SetBit("PN_Mixinghead_Send"); SetBit("PN_Mixinghead_Mixinghead{0}_DüseBypass{6}_Channel_Request"); SetBit("PN_Mixinghead_Mixinghead{0}_DüseBypass{6}_Zeiten_Request")
   "PN_Mixinghead_Mixinghead{0}_DüseBypass{6}_Active" : Bool = PLC PN_Mixinghead.Mixinghead[0].DüseBypass[6].Active AT %DB1006.DBX450.0, 1 s
      on ChangeValue: SetBit("PN_Mixinghead_Send"); SetBit("PN_Mixinghead_Mixinghead{0}_DüseBypass{6}_Channel_Request"); SetBit("PN_Mixinghead_Mixinghead{0}_DüseBypass{6}_Zeiten_Request")
   "PN_Mixinghead_Mixinghead{0}_DüseBypass{6}_Channel_Request" : Bool = PLC PN_Mixinghead.Mixinghead[0].DüseBypass[6].Channel.Request AT %DB1006.DBX452.0, 1 s
   "PN_Mixinghead_Mixinghead{0}_DüseBypass{1}_Channel_Request" : Bool = PLC PN_Mixinghead.Mixinghead[0].DüseBypass[1].Channel.Request AT %DB1006.DBX282.0, 1 s
   "PN_Mixinghead_Mixinghead{0}_DüseBypass{1}_Zeiten_Request" : Bool = PLC PN_Mixinghead.Mixinghead[0].DüseBypass[1].Zeiten.Request AT %DB1006.DBX288.0, 1 s
   "PN_Mixinghead_Mixinghead{0}_DüseBypass{2}_Channel_Request" : Bool = PLC PN_Mixinghead.Mixinghead[0].DüseBypass[2].Channel.Request AT %DB1006.DBX316.0, 1 s
   "PN_Mixinghead_Mixinghead{0}_DüseBypass{2}_Zeiten_Request" : Bool = PLC PN_Mixinghead.Mixinghead[0].DüseBypass[2].Zeiten.Request AT %DB1006.DBX322.0, 1 s
   "PN_Mixinghead_Mixinghead{0}_DüseBypass{3}_Channel_Request" : Bool = PLC PN_Mixinghead.Mixinghead[0].DüseBypass[3].Channel.Request AT %DB1006.DBX350.0, 1 s
   "PN_Mixinghead_Mixinghead{0}_DüseBypass{3}_Zeiten_Request" : Bool = PLC PN_Mixinghead.Mixinghead[0].DüseBypass[3].Zeiten.Request AT %DB1006.DBX356.0, 1 s
   "PN_Mixinghead_Mixinghead{0}_DüseBypass{4}_Channel_Request" : Bool = PLC PN_Mixinghead.Mixinghead[0].DüseBypass[4].Channel.Request AT %DB1006.DBX384.0, 1 s
   "PN_Mixinghead_Mixinghead{0}_DüseBypass{4}_Zeiten_Request" : Bool = PLC PN_Mixinghead.Mixinghead[0].DüseBypass[4].Zeiten.Request AT %DB1006.DBX390.0, 1 s
   "PN_Mixinghead_Mixinghead{0}_DüseBypass{5}_Channel_Request" : Bool = PLC PN_Mixinghead.Mixinghead[0].DüseBypass[5].Channel.Request AT %DB1006.DBX418.0, 1 s
   "PN_Mixinghead_Mixinghead{0}_DüseBypass{5}_Zeiten_Request" : Bool = PLC PN_Mixinghead.Mixinghead[0].DüseBypass[5].Zeiten.Request AT %DB1006.DBX424.0, 1 s
   "PN_Mixinghead_Mixinghead{0}_DüseBypass{1}_Visualisierung_OutputForNozzle" : Byte = PLC PN_Mixinghead.Mixinghead[0].DüseBypass[1].Visualisierung.OutputForNozzle AT %DB1006.DBB306, 1 s
      on ChangeValue: SetBit("PN_Mixinghead_Send"); SetBit("PN_Mixinghead_Mixinghead{0}_DüseBypass{1}_Channel_Request")
   "PN_Mixinghead_Mixinghead{0}_DüseBypass{1}_Visualisierung_PolarityNozzle" : Byte = PLC PN_Mixinghead.Mixinghead[0].DüseBypass[1].Visualisierung.PolarityNozzle AT %DB1006.DBB307, 1 s
      on ChangeValue: SetBit("PN_Mixinghead_Send"); SetBit("PN_Mixinghead_Mixinghead{0}_DüseBypass{1}_Channel_Request")
   "PN_Mixinghead_Mixinghead{0}_DüseBypass{1}_Visualisierung_OutputForBypass" : Byte = PLC PN_Mixinghead.Mixinghead[0].DüseBypass[1].Visualisierung.OutputForBypass AT %DB1006.DBB308, 1 s
      on ChangeValue: SetBit("PN_Mixinghead_Send"); SetBit("PN_Mixinghead_Mixinghead{0}_DüseBypass{1}_Channel_Request")
   "PN_Mixinghead_Mixinghead{0}_DüseBypass{1}_Visualisierung_PolarityBypass" : Byte = PLC PN_Mixinghead.Mixinghead[0].DüseBypass[1].Visualisierung.PolarityBypass AT %DB1006.DBB309, 1 s
      on ChangeValue: SetBit("PN_Mixinghead_Send"); SetBit("PN_Mixinghead_Mixinghead{0}_DüseBypass{1}_Channel_Request")
   "PN_Mixinghead_Mixinghead{0}_DüseBypass{1}_Visualisierung_MHChannel" : Byte = PLC PN_Mixinghead.Mixinghead[0].DüseBypass[1].Visualisierung.MHChannel AT %DB1006.DBB310, 1 s
      on ChangeValue: SetBit("PN_Mixinghead_Send"); SetBit("PN_Mixinghead_Mixinghead{0}_DüseBypass{1}_Channel_Request")
   "PN_Mixinghead_Mixinghead{0}_DüseBypass{2}_Visualisierung_OutputForNozzle" : Byte = PLC PN_Mixinghead.Mixinghead[0].DüseBypass[2].Visualisierung.OutputForNozzle AT %DB1006.DBB340, 1 s
      on ChangeValue: SetBit("PN_Mixinghead_Send"); SetBit("PN_Mixinghead_Mixinghead{0}_DüseBypass{2}_Channel_Request")
   "PN_Mixinghead_Mixinghead{0}_DüseBypass{2}_Visualisierung_PolarityNozzle" : Byte = PLC PN_Mixinghead.Mixinghead[0].DüseBypass[2].Visualisierung.PolarityNozzle AT %DB1006.DBB341, 1 s
      on ChangeValue: SetBit("PN_Mixinghead_Send"); SetBit("PN_Mixinghead_Mixinghead{0}_DüseBypass{2}_Channel_Request")
   "PN_Mixinghead_Mixinghead{0}_DüseBypass{2}_Visualisierung_OutputForBypass" : Byte = PLC PN_Mixinghead.Mixinghead[0].DüseBypass[2].Visualisierung.OutputForBypass AT %DB1006.DBB342, 1 s
      on ChangeValue: SetBit("PN_Mixinghead_Send"); SetBit("PN_Mixinghead_Mixinghead{0}_DüseBypass{2}_Channel_Request")
   "PN_Mixinghead_Mixinghead{0}_DüseBypass{2}_Visualisierung_PolarityBypass" : Byte = PLC PN_Mixinghead.Mixinghead[0].DüseBypass[2].Visualisierung.PolarityBypass AT %DB1006.DBB343, 1 s
      on ChangeValue: SetBit("PN_Mixinghead_Send"); SetBit("PN_Mixinghead_Mixinghead{0}_DüseBypass{2}_Channel_Request")
   "PN_Mixinghead_Mixinghead{0}_DüseBypass{2}_Visualisierung_MHChannel" : Byte = PLC PN_Mixinghead.Mixinghead[0].DüseBypass[2].Visualisierung.MHChannel AT %DB1006.DBB344, 1 s
      on ChangeValue: SetBit("PN_Mixinghead_Send"); SetBit("PN_Mixinghead_Mixinghead{0}_DüseBypass{2}_Channel_Request")
   "PN_Mixinghead_Mixinghead{0}_DüseBypass{3}_Visualisierung_OutputForNozzle" : Byte = PLC PN_Mixinghead.Mixinghead[0].DüseBypass[3].Visualisierung.OutputForNozzle AT %DB1006.DBB374, 1 s
      on ChangeValue: SetBit("PN_Mixinghead_Send"); SetBit("PN_Mixinghead_Mixinghead{0}_DüseBypass{3}_Channel_Request")
   "PN_Mixinghead_Mixinghead{0}_DüseBypass{3}_Visualisierung_PolarityNozzle" : Byte = PLC PN_Mixinghead.Mixinghead[0].DüseBypass[3].Visualisierung.PolarityNozzle AT %DB1006.DBB375, 1 s
      on ChangeValue: SetBit("PN_Mixinghead_Send"); SetBit("PN_Mixinghead_Mixinghead{0}_DüseBypass{3}_Channel_Request")
   "PN_Mixinghead_Mixinghead{0}_DüseBypass{3}_Visualisierung_OutputForBypass" : Byte = PLC PN_Mixinghead.Mixinghead[0].DüseBypass[3].Visualisierung.OutputForBypass AT %DB1006.DBB376, 1 s
      on ChangeValue: SetBit("PN_Mixinghead_Send"); SetBit("PN_Mixinghead_Mixinghead{0}_DüseBypass{3}_Channel_Request")
   "PN_Mixinghead_Mixinghead{0}_DüseBypass{3}_Visualisierung_PolarityBypass" : Byte = PLC PN_Mixinghead.Mixinghead[0].DüseBypass[3].Visualisierung.PolarityBypass AT %DB1006.DBB377, 1 s
      on ChangeValue: SetBit("PN_Mixinghead_Send"); SetBit("PN_Mixinghead_Mixinghead{0}_DüseBypass{3}_Channel_Request")
   "PN_Mixinghead_Mixinghead{0}_DüseBypass{3}_Visualisierung_MHChannel" : Byte = PLC PN_Mixinghead.Mixinghead[0].DüseBypass[3].Visualisierung.MHChannel AT %DB1006.DBB378, 1 s
      on ChangeValue: SetBit("PN_Mixinghead_Send"); SetBit("PN_Mixinghead_Mixinghead{0}_DüseBypass{3}_Channel_Request")
   "PN_Mixinghead_Mixinghead{0}_DüseBypass{4}_Visualisierung_OutputForNozzle" : Byte = PLC PN_Mixinghead.Mixinghead[0].DüseBypass[4].Visualisierung.OutputForNozzle AT %DB1006.DBB408, 1 s
      on ChangeValue: SetBit("PN_Mixinghead_Send"); SetBit("PN_Mixinghead_Mixinghead{0}_DüseBypass{4}_Channel_Request")
   "PN_Mixinghead_Mixinghead{0}_DüseBypass{4}_Visualisierung_PolarityNozzle" : Byte = PLC PN_Mixinghead.Mixinghead[0].DüseBypass[4].Visualisierung.PolarityNozzle AT %DB1006.DBB409, 1 s
      on ChangeValue: SetBit("PN_Mixinghead_Send"); SetBit("PN_Mixinghead_Mixinghead{0}_DüseBypass{4}_Channel_Request")
   "PN_Mixinghead_Mixinghead{0}_DüseBypass{4}_Visualisierung_OutputForBypass" : Byte = PLC PN_Mixinghead.Mixinghead[0].DüseBypass[4].Visualisierung.OutputForBypass AT %DB1006.DBB410, 1 s
      on ChangeValue: SetBit("PN_Mixinghead_Send"); SetBit("PN_Mixinghead_Mixinghead{0}_DüseBypass{4}_Channel_Request")
   "PN_Mixinghead_Mixinghead{0}_DüseBypass{4}_Visualisierung_PolarityBypass" : Byte = PLC PN_Mixinghead.Mixinghead[0].DüseBypass[4].Visualisierung.PolarityBypass AT %DB1006.DBB411, 1 s
      on ChangeValue: SetBit("PN_Mixinghead_Send"); SetBit("PN_Mixinghead_Mixinghead{0}_DüseBypass{4}_Channel_Request")
   "PN_Mixinghead_Mixinghead{0}_DüseBypass{4}_Visualisierung_MHChannel" : Byte = PLC PN_Mixinghead.Mixinghead[0].DüseBypass[4].Visualisierung.MHChannel AT %DB1006.DBB412, 1 s
      on ChangeValue: SetBit("PN_Mixinghead_Send"); SetBit("PN_Mixinghead_Mixinghead{0}_DüseBypass{4}_Channel_Request")
   "PN_Mixinghead_Mixinghead{0}_DüseBypass{5}_Visualisierung_OutputForNozzle" : Byte = PLC PN_Mixinghead.Mixinghead[0].DüseBypass[5].Visualisierung.OutputForNozzle AT %DB1006.DBB442, 1 s
      on ChangeValue: SetBit("PN_Mixinghead_Send"); SetBit("PN_Mixinghead_Mixinghead{0}_DüseBypass{5}_Channel_Request")
   "PN_Mixinghead_Mixinghead{0}_DüseBypass{5}_Visualisierung_PolarityNozzle" : Byte = PLC PN_Mixinghead.Mixinghead[0].DüseBypass[5].Visualisierung.PolarityNozzle AT %DB1006.DBB443, 1 s
      on ChangeValue: SetBit("PN_Mixinghead_Send"); SetBit("PN_Mixinghead_Mixinghead{0}_DüseBypass{5}_Channel_Request")
   "PN_Mixinghead_Mixinghead{0}_DüseBypass{5}_Visualisierung_OutputForBypass" : Byte = PLC PN_Mixinghead.Mixinghead[0].DüseBypass[5].Visualisierung.OutputForBypass AT %DB1006.DBB444, 1 s
      on ChangeValue: SetBit("PN_Mixinghead_Send"); SetBit("PN_Mixinghead_Mixinghead{0}_DüseBypass{5}_Channel_Request")
   "PN_Mixinghead_Mixinghead{0}_DüseBypass{5}_Visualisierung_PolarityBypass" : Byte = PLC PN_Mixinghead.Mixinghead[0].DüseBypass[5].Visualisierung.PolarityBypass AT %DB1006.DBB445, 1 s
      on ChangeValue: SetBit("PN_Mixinghead_Send"); SetBit("PN_Mixinghead_Mixinghead{0}_DüseBypass{5}_Channel_Request")
   "PN_Mixinghead_Mixinghead{0}_DüseBypass{5}_Visualisierung_MHChannel" : Byte = PLC PN_Mixinghead.Mixinghead[0].DüseBypass[5].Visualisierung.MHChannel AT %DB1006.DBB446, 1 s
      on ChangeValue: SetBit("PN_Mixinghead_Send"); SetBit("PN_Mixinghead_Mixinghead{0}_DüseBypass{5}_Channel_Request")
   "PN_Mixinghead_Mixinghead{0}_DüseBypass{6}_Visualisierung_OutputForNozzle" : Byte = PLC PN_Mixinghead.Mixinghead[0].DüseBypass[6].Visualisierung.OutputForNozzle AT %DB1006.DBB476, 1 s
      on ChangeValue: SetBit("PN_Mixinghead_Mixinghead{0}_DüseBypass{6}_Channel_Request"); SetBit("PN_Mixinghead_Send")
   "PN_Mixinghead_Mixinghead{0}_DüseBypass{6}_Visualisierung_PolarityNozzle" : Byte = PLC PN_Mixinghead.Mixinghead[0].DüseBypass[6].Visualisierung.PolarityNozzle AT %DB1006.DBB477, 1 s
      on ChangeValue: SetBit("PN_Mixinghead_Mixinghead{0}_DüseBypass{6}_Channel_Request"); SetBit("PN_Mixinghead_Send")
   "PN_Mixinghead_Mixinghead{0}_DüseBypass{6}_Visualisierung_OutputForBypass" : Byte = PLC PN_Mixinghead.Mixinghead[0].DüseBypass[6].Visualisierung.OutputForBypass AT %DB1006.DBB478, 1 s
      on ChangeValue: SetBit("PN_Mixinghead_Mixinghead{0}_DüseBypass{6}_Channel_Request"); SetBit("PN_Mixinghead_Send")
   "PN_Mixinghead_Mixinghead{0}_DüseBypass{6}_Visualisierung_PolarityBypass" : Byte = PLC PN_Mixinghead.Mixinghead[0].DüseBypass[6].Visualisierung.PolarityBypass AT %DB1006.DBB479, 1 s
      on ChangeValue: SetBit("PN_Mixinghead_Mixinghead{0}_DüseBypass{6}_Channel_Request"); SetBit("PN_Mixinghead_Send")
   "PN_Mixinghead_Mixinghead{0}_DüseBypass{6}_Visualisierung_MHChannel" : Byte = PLC PN_Mixinghead.Mixinghead[0].DüseBypass[6].Visualisierung.MHChannel AT %DB1006.DBB480, 1 s
      on ChangeValue: SetBit("PN_Mixinghead_Mixinghead{0}_DüseBypass{6}_Channel_Request"); SetBit("PN_Mixinghead_Send")
   "PN_Mixinghead_Mixinghead{0}_DüseBypass{1}_Zeiten_Data_ÜberlappungD_B" : Real = PLC PN_Mixinghead.Mixinghead[0].DüseBypass[1].Zeiten.Data.ÜberlappungD_B AT %DB1006.DBD290, 1 s
      on ChangeValue: SetBit("PN_Mixinghead_Send"); SetBit("PN_Mixinghead_Mixinghead{0}_DüseBypass{1}_Zeiten_Request")
   "PN_Mixinghead_Mixinghead{0}_DüseBypass{1}_Zeiten_Data_ÜberlappungB_D" : Real = PLC PN_Mixinghead.Mixinghead[0].DüseBypass[1].Zeiten.Data.ÜberlappungB_D AT %DB1006.DBD294, 1 s
      on ChangeValue: SetBit("PN_Mixinghead_Send"); SetBit("PN_Mixinghead_Mixinghead{0}_DüseBypass{1}_Zeiten_Request")
   "PN_Mixinghead_Mixinghead{0}_DüseBypass{1}_Zeiten_Data_VerzögerungSchussstart" : Real = PLC PN_Mixinghead.Mixinghead[0].DüseBypass[1].Zeiten.Data.VerzögerungSchussstart AT %DB1006.DBD298, 1 s
      on ChangeValue: SetBit("PN_Mixinghead_Send"); SetBit("PN_Mixinghead_Mixinghead{0}_DüseBypass{1}_Zeiten_Request")
   "PN_Mixinghead_Mixinghead{0}_DüseBypass{1}_Zeiten_Data_VerzögerungSchussende" : Real = PLC PN_Mixinghead.Mixinghead[0].DüseBypass[1].Zeiten.Data.VerzögerungSchussende AT %DB1006.DBD302, 1 s
      on ChangeValue: SetBit("PN_Mixinghead_Send"); SetBit("PN_Mixinghead_Mixinghead{0}_DüseBypass{1}_Zeiten_Request")
   "PN_Mixinghead_Mixinghead{0}_DüseBypass{2}_Zeiten_Data_ÜberlappungD_B" : Real = PLC PN_Mixinghead.Mixinghead[0].DüseBypass[2].Zeiten.Data.ÜberlappungD_B AT %DB1006.DBD324, 1 s
      on ChangeValue: SetBit("PN_Mixinghead_Send"); SetBit("PN_Mixinghead_Mixinghead{0}_DüseBypass{2}_Zeiten_Request")
   "PN_Mixinghead_Mixinghead{0}_DüseBypass{2}_Zeiten_Data_ÜberlappungB_D" : Real = PLC PN_Mixinghead.Mixinghead[0].DüseBypass[2].Zeiten.Data.ÜberlappungB_D AT %DB1006.DBD328, 1 s
      on ChangeValue: SetBit("PN_Mixinghead_Send"); SetBit("PN_Mixinghead_Mixinghead{0}_DüseBypass{2}_Zeiten_Request")
   "PN_Mixinghead_Mixinghead{0}_DüseBypass{2}_Zeiten_Data_VerzögerungSchussstart" : Real = PLC PN_Mixinghead.Mixinghead[0].DüseBypass[2].Zeiten.Data.VerzögerungSchussstart AT %DB1006.DBD332, 1 s
      on ChangeValue: SetBit("PN_Mixinghead_Send"); SetBit("PN_Mixinghead_Mixinghead{0}_DüseBypass{2}_Zeiten_Request")
   "PN_Mixinghead_Mixinghead{0}_DüseBypass{2}_Zeiten_Data_VerzögerungSchussende" : Real = PLC PN_Mixinghead.Mixinghead[0].DüseBypass[2].Zeiten.Data.VerzögerungSchussende AT %DB1006.DBD336, 1 s
      on ChangeValue: SetBit("PN_Mixinghead_Send"); SetBit("PN_Mixinghead_Mixinghead{0}_DüseBypass{2}_Zeiten_Request")
   "PN_Mixinghead_Mixinghead{0}_DüseBypass{3}_Zeiten_Data_ÜberlappungD_B" : Real = PLC PN_Mixinghead.Mixinghead[0].DüseBypass[3].Zeiten.Data.ÜberlappungD_B AT %DB1006.DBD358, 1 s
      on ChangeValue: SetBit("PN_Mixinghead_Send"); SetBit("PN_Mixinghead_Mixinghead{0}_DüseBypass{3}_Zeiten_Request")
   "PN_Mixinghead_Mixinghead{0}_DüseBypass{3}_Zeiten_Data_ÜberlappungB_D" : Real = PLC PN_Mixinghead.Mixinghead[0].DüseBypass[3].Zeiten.Data.ÜberlappungB_D AT %DB1006.DBD362, 1 s
      on ChangeValue: SetBit("PN_Mixinghead_Send"); SetBit("PN_Mixinghead_Mixinghead{0}_DüseBypass{3}_Zeiten_Request")
   "PN_Mixinghead_Mixinghead{0}_DüseBypass{3}_Zeiten_Data_VerzögerungSchussstart" : Real = PLC PN_Mixinghead.Mixinghead[0].DüseBypass[3].Zeiten.Data.VerzögerungSchussstart AT %DB1006.DBD366, 1 s
      on ChangeValue: SetBit("PN_Mixinghead_Send"); SetBit("PN_Mixinghead_Mixinghead{0}_DüseBypass{3}_Zeiten_Request")
   "PN_Mixinghead_Mixinghead{0}_DüseBypass{3}_Zeiten_Data_VerzögerungSchussende" : Real = PLC PN_Mixinghead.Mixinghead[0].DüseBypass[3].Zeiten.Data.VerzögerungSchussende AT %DB1006.DBD370, 1 s
      on ChangeValue: SetBit("PN_Mixinghead_Send"); SetBit("PN_Mixinghead_Mixinghead{0}_DüseBypass{3}_Zeiten_Request")